REGION Network 15
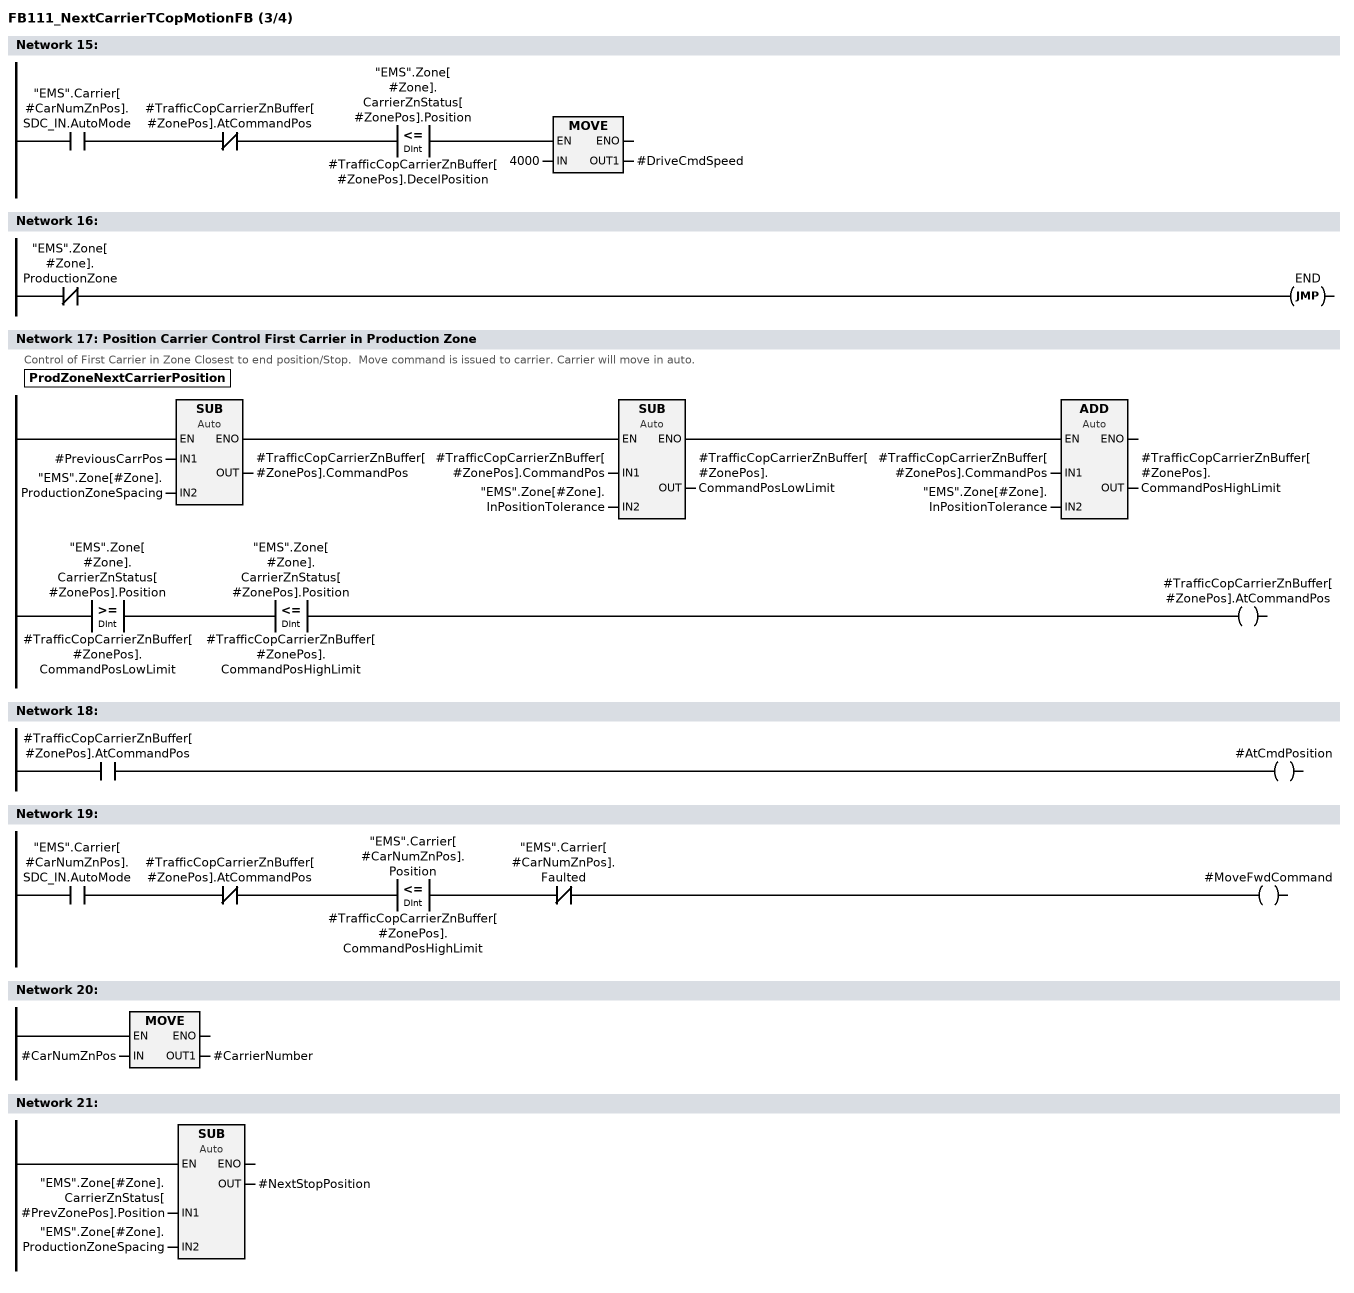
   RUNG wire#powerrail
      Contact( "EMS".Carrier[#CarNumZnPos].SDC_IN.AutoMode )
      I_Contact( #TrafficCopCarrierZnBuffer[#ZonePos].AtCommandPos )
      { S7_Templates := "SrcType := DInt" } LE_Contact(in1 := "EMS".Zone[#Zone].CarrierZnStatus[#ZonePos].Position, in2 := #TrafficCopCarrierZnBuffer[#ZonePos].DecelPosition)
      Move(in := 4000, out1 => #DriveCmdSpeed)
   END_RUNG
   // the same network as SCL:
   IF "EMS".Carrier[#CarNumZnPos].SDC_IN.AutoMode AND NOT #TrafficCopCarrierZnBuffer[#ZonePos].AtCommandPos AND ("EMS".Zone[#Zone].CarrierZnStatus[#ZonePos].Position <= #TrafficCopCarrierZnBuffer[#ZonePos].DecelPosition) THEN
       #DriveCmdSpeed := 4000;
   END_IF;
END_REGION

REGION Network 16
   RUNG wire#powerrail
      I_Contact( "EMS".Zone[#Zone].ProductionZone )
      JumpCoil( END )
   END_RUNG
   // the same network as SCL:
   IF NOT "EMS".Zone[#Zone].ProductionZone THEN GOTO END; END_IF;
END_REGION

REGION Network 17: Position Carrier Control First Carrier in Production Zone
   // Control of First Carrier in Zone Closest to end position/Stop.  Move command is issued to carrier. Carrier will move in auto.
   Label( ProdZoneNextCarrierPosition )
   RUNG wire#powerrail
      Sub(in1 := #PreviousCarrPos, in2 := "EMS".Zone[#Zone].ProductionZoneSpacing, out => #TrafficCopCarrierZnBuffer[#ZonePos].CommandPos)
      Sub(in1 := #TrafficCopCarrierZnBuffer[#ZonePos].CommandPos, in2 := "EMS".Zone[#Zone].InPositionTolerance, out => #TrafficCopCarrierZnBuffer[#ZonePos].CommandPosLowLimit)
      Add(in1 := #TrafficCopCarrierZnBuffer[#ZonePos].CommandPos, in2 := "EMS".Zone[#Zone].InPositionTolerance, out => #TrafficCopCarrierZnBuffer[#ZonePos].CommandPosHighLimit)
   END_RUNG
   RUNG wire#powerrail
      { S7_Templates := "SrcType := DInt" } GE_Contact(in1 := "EMS".Zone[#Zone].CarrierZnStatus[#ZonePos].Position, in2 := #TrafficCopCarrierZnBuffer[#ZonePos].CommandPosLowLimit)
      { S7_Templates := "SrcType := DInt" } LE_Contact(in1 := "EMS".Zone[#Zone].CarrierZnStatus[#ZonePos].Position, in2 := #TrafficCopCarrierZnBuffer[#ZonePos].CommandPosHighLimit)
      Coil( #TrafficCopCarrierZnBuffer[#ZonePos].AtCommandPos )
   END_RUNG
   // the same network as SCL:
   ProdZoneNextCarrierPosition:
   #TrafficCopCarrierZnBuffer[#ZonePos].CommandPos := #PreviousCarrPos - "EMS".Zone[#Zone].ProductionZoneSpacing;
   #TrafficCopCarrierZnBuffer[#ZonePos].CommandPosLowLimit := #TrafficCopCarrierZnBuffer[#ZonePos].CommandPos - "EMS".Zone[#Zone].InPositionTolerance;
   #TrafficCopCarrierZnBuffer[#ZonePos].CommandPosHighLimit := #TrafficCopCarrierZnBuffer[#ZonePos].CommandPos + "EMS".Zone[#Zone].InPositionTolerance;
   #TrafficCopCarrierZnBuffer[#ZonePos].AtCommandPos := ("EMS".Zone[#Zone].CarrierZnStatus[#ZonePos].Position >= #TrafficCopCarrierZnBuffer[#ZonePos].CommandPosLowLimit) AND ("EMS".Zone[#Zone].CarrierZnStatus[#ZonePos].Position <= #TrafficCopCarrierZnBuffer[#ZonePos].CommandPosHighLimit);
END_REGION

REGION Network 18
   RUNG wire#powerrail
      Contact( #TrafficCopCarrierZnBuffer[#ZonePos].AtCommandPos )
      Coil( #AtCmdPosition )
   END_RUNG
   // the same network as SCL:
   #AtCmdPosition := #TrafficCopCarrierZnBuffer[#ZonePos].AtCommandPos;
END_REGION

REGION Network 19
   RUNG wire#powerrail
      Contact( "EMS".Carrier[#CarNumZnPos].SDC_IN.AutoMode )
      I_Contact( #TrafficCopCarrierZnBuffer[#ZonePos].AtCommandPos )
      { S7_Templates := "SrcType := DInt" } LE_Contact(in1 := "EMS".Carrier[#CarNumZnPos].Position, in2 := #TrafficCopCarrierZnBuffer[#ZonePos].CommandPosHighLimit)
      I_Contact( "EMS".Carrier[#CarNumZnPos].Faulted )
      Coil( #MoveFwdCommand )
   END_RUNG
   // the same network as SCL:
   #MoveFwdCommand := "EMS".Carrier[#CarNumZnPos].SDC_IN.AutoMode AND NOT #TrafficCopCarrierZnBuffer[#ZonePos].AtCommandPos AND ("EMS".Carrier[#CarNumZnPos].Position <= #TrafficCopCarrierZnBuffer[#ZonePos].CommandPosHighLimit) AND NOT "EMS".Carrier[#CarNumZnPos].Faulted;
END_REGION

REGION Network 20
   RUNG wire#powerrail
      Move(in := #CarNumZnPos, out1 => #CarrierNumber)
   END_RUNG
   // the same network as SCL:
   #CarrierNumber := #CarNumZnPos;
END_REGION

REGION Network 21
   RUNG wire#powerrail
      Sub(in1 := "EMS".Zone[#Zone].CarrierZnStatus[#PrevZonePos].Position, in2 := "EMS".Zone[#Zone].ProductionZoneSpacing, out => #NextStopPosition)
   END_RUNG
   // the same network as SCL:
   #NextStopPosition := "EMS".Zone[#Zone].CarrierZnStatus[#PrevZonePos].Position - "EMS".Zone[#Zone].ProductionZoneSpacing;
END_REGION

REGION Network 22
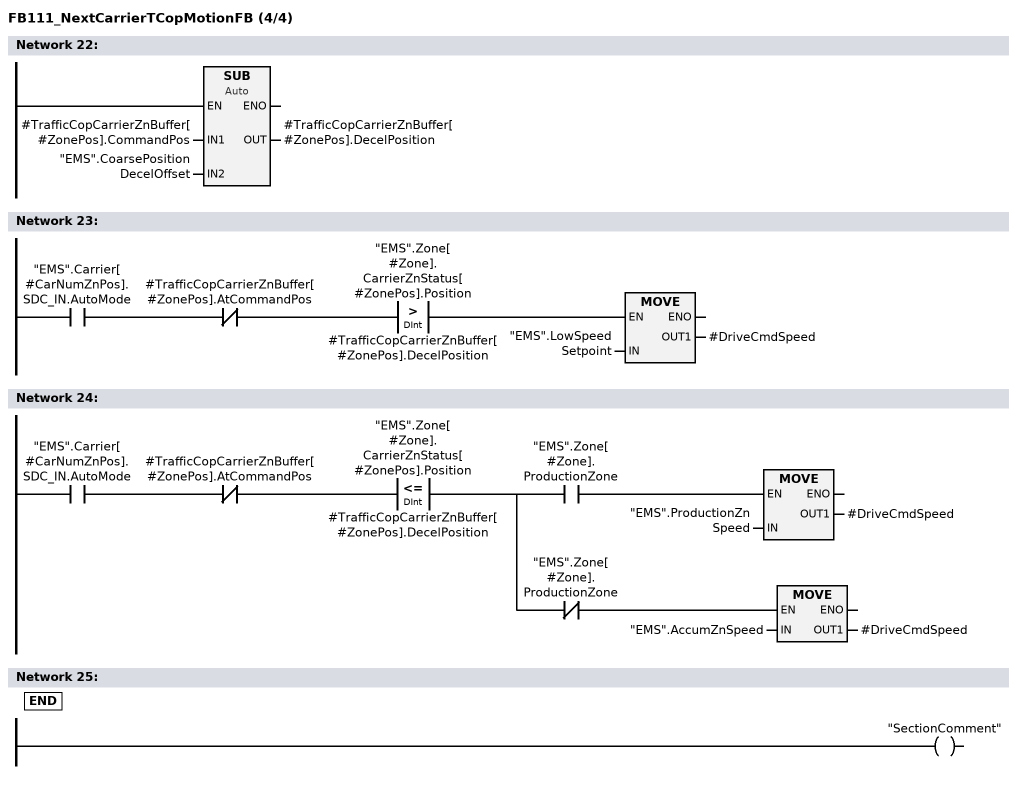
   RUNG wire#powerrail
      Sub(in1 := #TrafficCopCarrierZnBuffer[#ZonePos].CommandPos, in2 := "EMS".CoarsePositionDecelOffset, out => #TrafficCopCarrierZnBuffer[#ZonePos].DecelPosition)
   END_RUNG
   // the same network as SCL:
   #TrafficCopCarrierZnBuffer[#ZonePos].DecelPosition := #TrafficCopCarrierZnBuffer[#ZonePos].CommandPos - "EMS".CoarsePositionDecelOffset;
END_REGION

REGION Network 23
   RUNG wire#powerrail
      Contact( "EMS".Carrier[#CarNumZnPos].SDC_IN.AutoMode )
      I_Contact( #TrafficCopCarrierZnBuffer[#ZonePos].AtCommandPos )
      { S7_Templates := "SrcType := DInt" } GT_Contact(in1 := "EMS".Zone[#Zone].CarrierZnStatus[#ZonePos].Position, in2 := #TrafficCopCarrierZnBuffer[#ZonePos].DecelPosition)
      Move(in := "EMS".LowSpeedSetpoint, out1 => #DriveCmdSpeed)
   END_RUNG
   // the same network as SCL:
   IF "EMS".Carrier[#CarNumZnPos].SDC_IN.AutoMode AND NOT #TrafficCopCarrierZnBuffer[#ZonePos].AtCommandPos AND ("EMS".Zone[#Zone].CarrierZnStatus[#ZonePos].Position > #TrafficCopCarrierZnBuffer[#ZonePos].DecelPosition) THEN
       #DriveCmdSpeed := "EMS".LowSpeedSetpoint;
   END_IF;
END_REGION

REGION Network 24
   RUNG wire#powerrail
      Contact( "EMS".Carrier[#CarNumZnPos].SDC_IN.AutoMode )
      I_Contact( #TrafficCopCarrierZnBuffer[#ZonePos].AtCommandPos )
      { S7_Templates := "SrcType := DInt" } LE_Contact(in1 := "EMS".Zone[#Zone].CarrierZnStatus[#ZonePos].Position, in2 := #TrafficCopCarrierZnBuffer[#ZonePos].DecelPosition)
      wire#w1
      Contact( "EMS".Zone[#Zone].ProductionZone )
      Move(in := "EMS".ProductionZnSpeed, out1 => #DriveCmdSpeed)
   END_RUNG
   RUNG wire#w1
      I_Contact( "EMS".Zone[#Zone].ProductionZone )
      Move(in := "EMS".AccumZnSpeed, out1 => #DriveCmdSpeed)
   END_RUNG
   // the same network as SCL:
   #_w1 := "EMS".Carrier[#CarNumZnPos].SDC_IN.AutoMode AND NOT #TrafficCopCarrierZnBuffer[#ZonePos].AtCommandPos AND ("EMS".Zone[#Zone].CarrierZnStatus[#ZonePos].Position <= #TrafficCopCarrierZnBuffer[#ZonePos].DecelPosition);
   IF #_w1 AND "EMS".Zone[#Zone].ProductionZone THEN #DriveCmdSpeed := "EMS".ProductionZnSpeed; END_IF;
   IF #_w1 AND NOT "EMS".Zone[#Zone].ProductionZone THEN #DriveCmdSpeed := "EMS".AccumZnSpeed; END_IF;
END_REGION

REGION Network 25
   Label( END )
   RUNG wire#powerrail
      Coil( "SectionComment" )
   END_RUNG
   // the same network as SCL:
   END:
   "SectionComment" := TRUE;
END_REGION
END_FUNCTION_BLOCK

FUNCTION_BLOCK "FB112_Carrier"   // FB112, LAD
{ S7_Optimized_Access := 'TRUE' }
VERSION : 0.1
   VAR_INPUT
      Carrier : Int;
      EMS : "UDT_System";
      MoveFwd : Bool;
      SpeedSelect : Word;   // Speed Select 1=Slow 2=Normal
      CarrierFindArrayBufferiN : "UDT_Carrier";
      SDC_IN : "UDT_SDC_IN";
      DuplicateCarrierNumIn : Int;
      DuplicateCarrierFound : Bool;
      GapSpacingFault : Bool;
      FaultReset : Bool;
   END_VAR
   VAR_OUTPUT
      Zone : Int;
      ZonePos : Word;
      CarrierPositionEcho : DWord;
      CarrierNumberEcho : Word;
      DuplicateCarrierNumEcho : Word;
      CarrierNextStopPosEcho : Word;
      Faults : "UDT_SDCOutFaults";
      Faulted : Bool;
   END_VAR
   VAR
      CarrierMoveFwdSetup : Array[0..30] of Bool;
      MotionOffFaultTimer : IEC_TIMER;
      MotionOnFaultTimer : IEC_TIMER;
   END_VAR
BEGIN

REGION Network 1
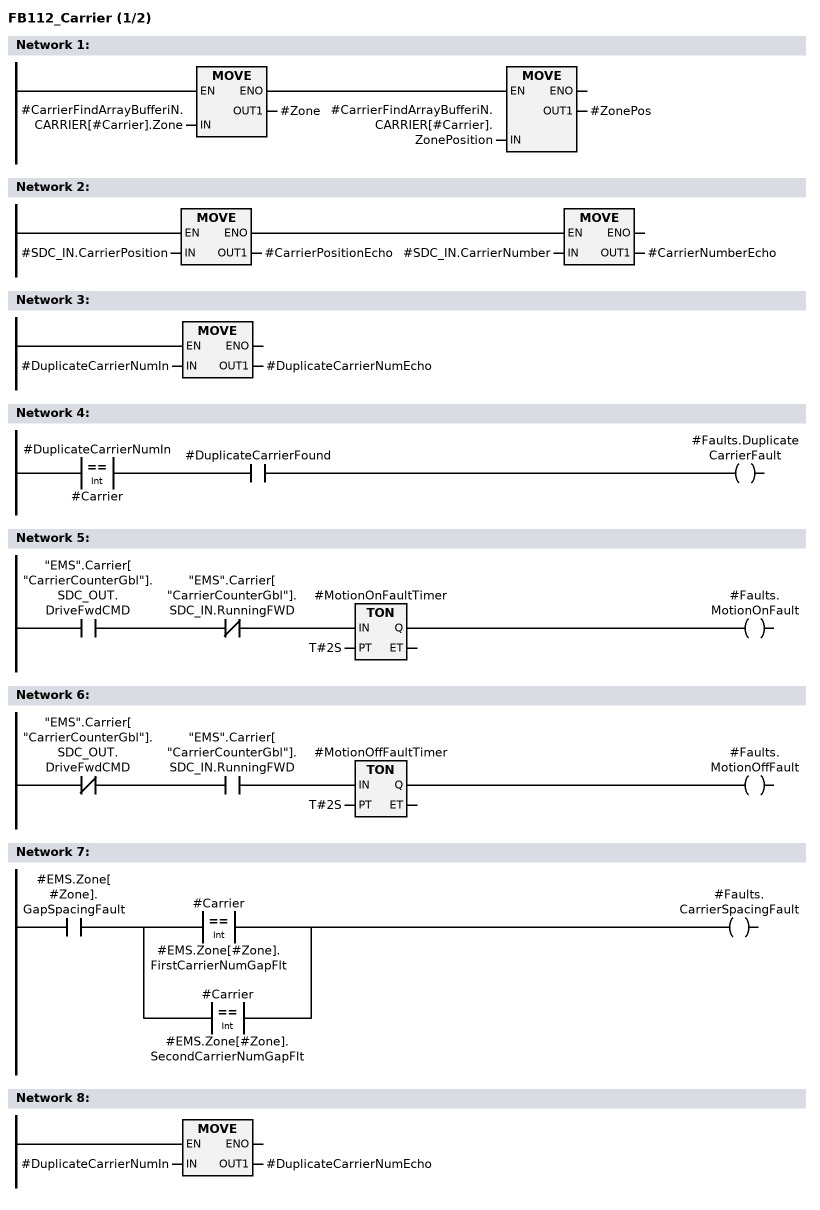
   RUNG wire#powerrail
      Move(in := #CarrierFindArrayBufferiN.CARRIER[#Carrier].Zone, out1 => #Zone)
      Move(in := #CarrierFindArrayBufferiN.CARRIER[#Carrier].ZonePosition, out1 => #ZonePos)
   END_RUNG
   // the same network as SCL:
   #Zone := #CarrierFindArrayBufferiN.CARRIER[#Carrier].Zone;
   #ZonePos := #CarrierFindArrayBufferiN.CARRIER[#Carrier].ZonePosition;
END_REGION

REGION Network 2
   RUNG wire#powerrail
      Move(in := #SDC_IN.CarrierPosition, out1 => #CarrierPositionEcho)
      Move(in := #SDC_IN.CarrierNumber, out1 => #CarrierNumberEcho)
   END_RUNG
   // the same network as SCL:
   #CarrierPositionEcho := #SDC_IN.CarrierPosition;
   #CarrierNumberEcho := #SDC_IN.CarrierNumber;
END_REGION

REGION Network 3
   RUNG wire#powerrail
      Move(in := #DuplicateCarrierNumIn, out1 => #DuplicateCarrierNumEcho)
   END_RUNG
   // the same network as SCL:
   #DuplicateCarrierNumEcho := #DuplicateCarrierNumIn;
END_REGION

REGION Network 4
   RUNG wire#powerrail
      { S7_Templates := "SrcType := Int" } EQ_Contact(in1 := #DuplicateCarrierNumIn, in2 := #Carrier)
      Contact( #DuplicateCarrierFound )
      Coil( #Faults.DuplicateCarrierFault )
   END_RUNG
   // the same network as SCL:
   #Faults.DuplicateCarrierFault := (#DuplicateCarrierNumIn = #Carrier) AND #DuplicateCarrierFound;
END_REGION

REGION Network 5
   #MotionOnFaultTimer.TON(IN := "EMS".Carrier["CarrierCounterGbl"].SDC_OUT.DriveFwdCMD AND NOT "EMS".Carrier["CarrierCounterGbl"].SDC_IN.RunningFWD,
                           PT := T#2S);
   #Faults.MotionOnFault := #MotionOnFaultTimer.Q;
END_REGION

REGION Network 6
   #MotionOffFaultTimer.TON(IN := NOT "EMS".Carrier["CarrierCounterGbl"].SDC_OUT.DriveFwdCMD AND "EMS".Carrier["CarrierCounterGbl"].SDC_IN.RunningFWD,
                           PT := T#2S);
   #Faults.MotionOffFault := #MotionOffFaultTimer.Q;
END_REGION

REGION Network 7
   RUNG wire#powerrail
      Contact( #EMS.Zone[#Zone].GapSpacingFault )
      wire#w1
      { S7_Templates := "SrcType := Int" } EQ_Contact(in1 := #Carrier, in2 := #EMS.Zone[#Zone].FirstCarrierNumGapFlt)
      wire#w2
      Coil( #Faults.CarrierSpacingFault )
   END_RUNG
   RUNG wire#w1
      { S7_Templates := "SrcType := Int" } EQ_Contact(in1 := #Carrier, in2 := #EMS.Zone[#Zone].SecondCarrierNumGapFlt)
   END_RUNG wire#w2
   // the same network as SCL:
   #Faults.CarrierSpacingFault := #EMS.Zone[#Zone].GapSpacingFault AND ((#Carrier = #EMS.Zone[#Zone].FirstCarrierNumGapFlt) OR (#Carrier = #EMS.Zone[#Zone].SecondCarrierNumGapFlt));
END_REGION

REGION Network 8
   RUNG wire#powerrail
      Move(in := #DuplicateCarrierNumIn, out1 => #DuplicateCarrierNumEcho)
   END_RUNG
   // the same network as SCL:
   #DuplicateCarrierNumEcho := #DuplicateCarrierNumIn;
END_REGION

REGION Network 9
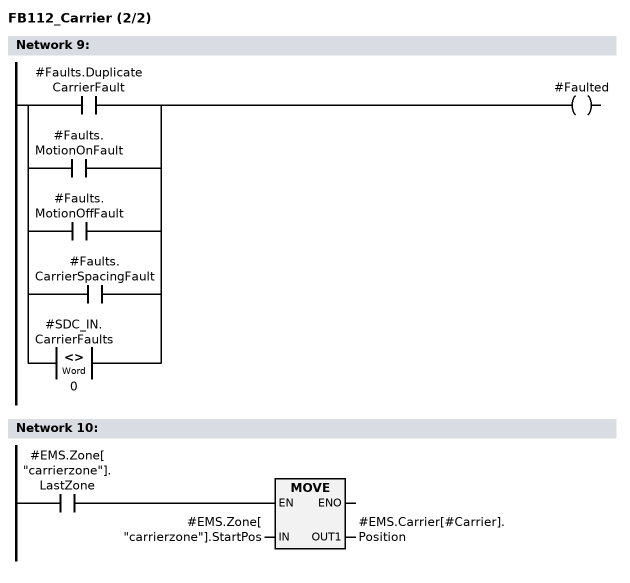
   RUNG wire#powerrail
      Contact( #Faults.DuplicateCarrierFault )
      wire#w1
      Coil( #Faulted )
   END_RUNG
   RUNG wire#powerrail
      Contact( #Faults.MotionOnFault )
   END_RUNG wire#w1
   RUNG wire#powerrail
      Contact( #Faults.MotionOffFault )
   END_RUNG wire#w1
   RUNG wire#powerrail
      Contact( #Faults.CarrierSpacingFault )
   END_RUNG wire#w1
   RUNG wire#powerrail
      { S7_Templates := "SrcType := Word" } NE_Contact(in1 := #SDC_IN.CarrierFaults, in2 := 0)
   END_RUNG wire#w1
   // the same network as SCL:
   #Faulted := #Faults.DuplicateCarrierFault OR #Faults.MotionOnFault OR #Faults.MotionOffFault OR #Faults.CarrierSpacingFault OR (#SDC_IN.CarrierFaults <> 0);
END_REGION

REGION Network 10
   RUNG wire#powerrail
      Contact( #EMS.Zone["carrierzone"].LastZone )
      Move(in := #EMS.Zone["carrierzone"].StartPos, out1 => #EMS.Carrier[#Carrier].Position)
   END_RUNG
   // the same network as SCL:
   IF #EMS.Zone["carrierzone"].LastZone THEN
       #EMS.Carrier[#Carrier].Position := #EMS.Zone["carrierzone"].StartPos;
   END_IF;
END_REGION
END_FUNCTION_BLOCK

FUNCTION_BLOCK "FB113_CarrierTrafficCop"   // FB113, LAD
{ S7_Optimized_Access := 'TRUE' }
VERSION : 0.1
   VAR_INPUT
      CarrierNumber : Word;
      ZonePos : Word;
   END_VAR
BEGIN
END_FUNCTION_BLOCK

FUNCTION_BLOCK "FB115_FB_Zone"   // FB115, LAD
{ S7_Optimized_Access := 'FALSE' }
VERSION : 0.1
   VAR_INPUT
      Zone : Int;
      Description : String[10];
      LastZone : Bool;
      MaxCarriers : Int;
      StartPos : DWord;
      EndPos : DWord;
      NextZone : Word;   // If Zone numbering is non sequential Next Zone Nu
      PreviousZone : Word;   // If Zone numbering is non sequential Previous Zone Nu
      SpeedZone : Bool;
      SpeedZoneStart : DWord;
      SpeedZoneEnd : DWord;
      AccumZone : Bool;
      AccumZnSpacing : Word;
      ProductionZone : Bool := false;
      ProductZoneSpacing : Word;
      FinePosStopZone : Bool;
      FineInPosTolerance : Word;
      FinePositionDecelOffset : Word;
      CoarseInPosTolerance : Word;
      CoarsePositionDecelOffset : Word;
      NextCarrierClrHighSpeed : Word;
      StopControlFromEMS01 : "UDT_StopControlFromEMS01";
   END_VAR
   VAR_OUTPUT
      ZoneEcho : Word;
      LastZoneEcho : Bool;
      ZoneFull : Bool;
      ZoneLengthEcho : Word;
      DescriptionEcho : String[10];
      StartPosEcho : DWord;
      EndPosEcho : DWord;
      SpeedZoneEcho : Bool;
      SpeedZoneStartEcho : DWord;
      SpeedZoneEndEcho : DWord;
      AccumZoneEcho : Bool;
      AccumSpacingEcho : Word;
      ProductionZoneEcho : Bool;
      ProdZoneSpacingEcho : Word;
      CarrierInPosToleranceEcho : Word;
      NextCarrierClrHighSpeedEcho : Word;
      MaxCarriersEcho : Word;
      ClearToEnterEcho : Bool;
      ClearZoneStartEcho : Bool;
      ClearZoneEcho : Bool;
      ZoneCarrierStatsArray : Array[0..60] of "UDT_ZoneCarrierStatus";
      FinePosStopZoneEcho : Bool;
      FineInPosToleranceEcho : Word;
      FinePositionDecelEcho : Word;
      CoarsePositionDecelEcho : Word;
      CoarseInPosToleranceEcho : Word;
      PreviosZoneEcho : Word;
      NextZoneEcho : Word;
      CarrierAtStop : Bool;
      CarrierNumAtStop : Word;
      HMIZonePositionsEcho : Array[1..20] of "UDT_HMIZonePositions";
      ClearOfStopPos : DWord;
      StopStatusToEMS01 : "UDT_StopStatusToEMS01";
   END_VAR
   VAR_TEMP
      HMIZonePositions : Array[1..20] of "UDT_HMIZonePositions";
      carrierstatusdn : Bool;
      resettemp : Bool;
      resettemp2 : Bool;
      sortdonetemp : Bool;
      ZonePosSpacing : Word;
      ZoneLengthTemp : UDInt;
   END_VAR
BEGIN

REGION Network 1
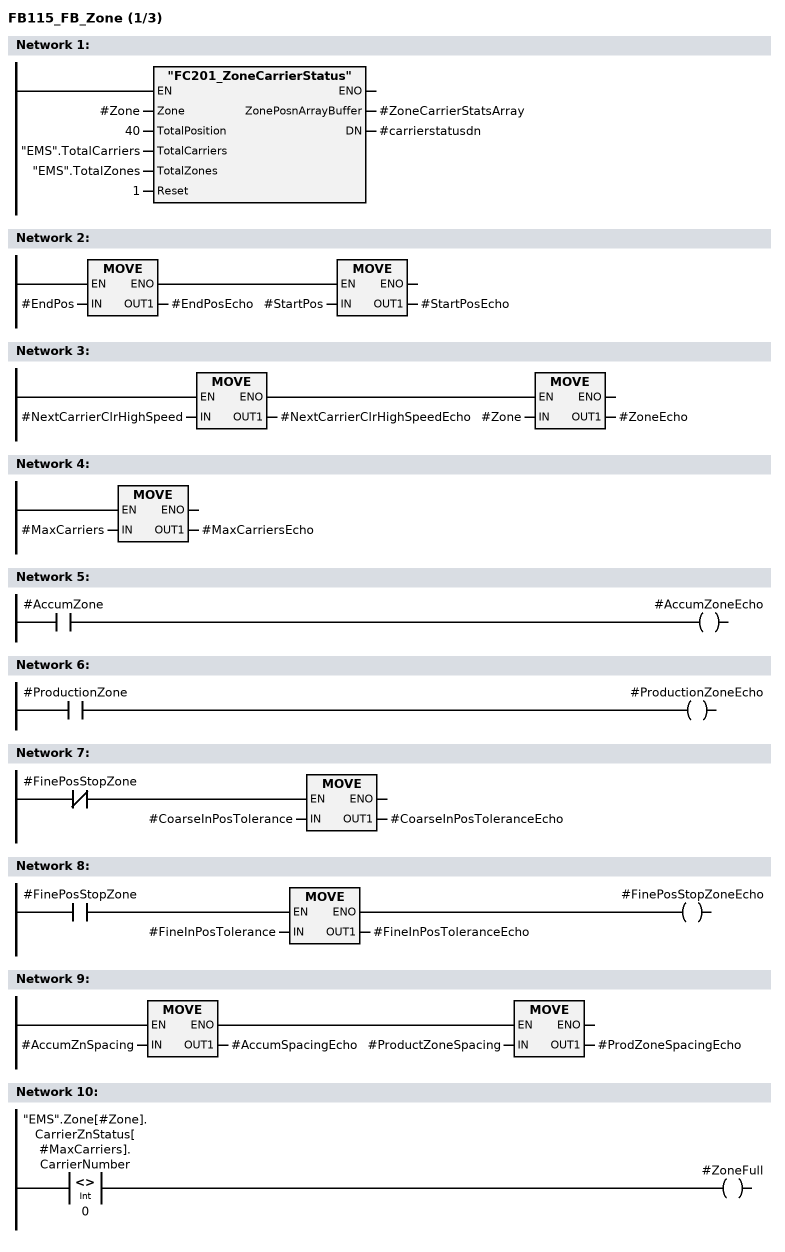
   RUNG wire#powerrail
      "FC201_ZoneCarrierStatus"(Zone := #Zone, TotalPosition := 40, TotalCarriers := "EMS".TotalCarriers, TotalZones := "EMS".TotalZones, Reset := 1, ZonePosnArrayBuffer => #ZoneCarrierStatsArray, DN => #carrierstatusdn)
   END_RUNG
   // the same network as SCL:
   "FC201_ZoneCarrierStatus"(Zone := #Zone,
                           TotalPosition := 40,
                           TotalCarriers := "EMS".TotalCarriers,
                           TotalZones := "EMS".TotalZones,
                           Reset := 1,
                           ZonePosnArrayBuffer => #ZoneCarrierStatsArray,
                           DN => #carrierstatusdn);
END_REGION

REGION Network 2
   RUNG wire#powerrail
      Move(in := #EndPos, out1 => #EndPosEcho)
      Move(in := #StartPos, out1 => #StartPosEcho)
   END_RUNG
   // the same network as SCL:
   #EndPosEcho := #EndPos;
   #StartPosEcho := #StartPos;
END_REGION

REGION Network 3
   RUNG wire#powerrail
      Move(in := #NextCarrierClrHighSpeed, out1 => #NextCarrierClrHighSpeedEcho)
      Move(in := #Zone, out1 => #ZoneEcho)
   END_RUNG
   // the same network as SCL:
   #NextCarrierClrHighSpeedEcho := #NextCarrierClrHighSpeed;
   #ZoneEcho := #Zone;
END_REGION

REGION Network 4
   RUNG wire#powerrail
      Move(in := #MaxCarriers, out1 => #MaxCarriersEcho)
   END_RUNG
   // the same network as SCL:
   #MaxCarriersEcho := #MaxCarriers;
END_REGION

REGION Network 5
   RUNG wire#powerrail
      Contact( #AccumZone )
      Coil( #AccumZoneEcho )
   END_RUNG
   // the same network as SCL:
   #AccumZoneEcho := #AccumZone;
END_REGION

REGION Network 6
   RUNG wire#powerrail
      Contact( #ProductionZone )
      Coil( #ProductionZoneEcho )
   END_RUNG
   // the same network as SCL:
   #ProductionZoneEcho := #ProductionZone;
END_REGION

REGION Network 7
   RUNG wire#powerrail
      I_Contact( #FinePosStopZone )
      Move(in := #CoarseInPosTolerance, out1 => #CoarseInPosToleranceEcho)
   END_RUNG
   // the same network as SCL:
   IF NOT #FinePosStopZone THEN #CoarseInPosToleranceEcho := #CoarseInPosTolerance; END_IF;
END_REGION

REGION Network 8
   RUNG wire#powerrail
      Contact( #FinePosStopZone )
      Move(in := #FineInPosTolerance, out1 => #FineInPosToleranceEcho)
      Coil( #FinePosStopZoneEcho )
   END_RUNG
   // the same network as SCL:
   IF #FinePosStopZone THEN #FineInPosToleranceEcho := #FineInPosTolerance; END_IF;
   #FinePosStopZoneEcho := #FinePosStopZone;
END_REGION

REGION Network 9
   RUNG wire#powerrail
      Move(in := #AccumZnSpacing, out1 => #AccumSpacingEcho)
      Move(in := #ProductZoneSpacing, out1 => #ProdZoneSpacingEcho)
   END_RUNG
   // the same network as SCL:
   #AccumSpacingEcho := #AccumZnSpacing;
   #ProdZoneSpacingEcho := #ProductZoneSpacing;
END_REGION

REGION Network 10
   RUNG wire#powerrail
      { S7_Templates := "SrcType := Int" } NE_Contact(in1 := "EMS".Zone[#Zone].CarrierZnStatus[#MaxCarriers].CarrierNumber, in2 := 0)
      Coil( #ZoneFull )
   END_RUNG
   // the same network as SCL:
   #ZoneFull := "EMS".Zone[#Zone].CarrierZnStatus[#MaxCarriers].CarrierNumber <> 0;
END_REGION

REGION Network 11
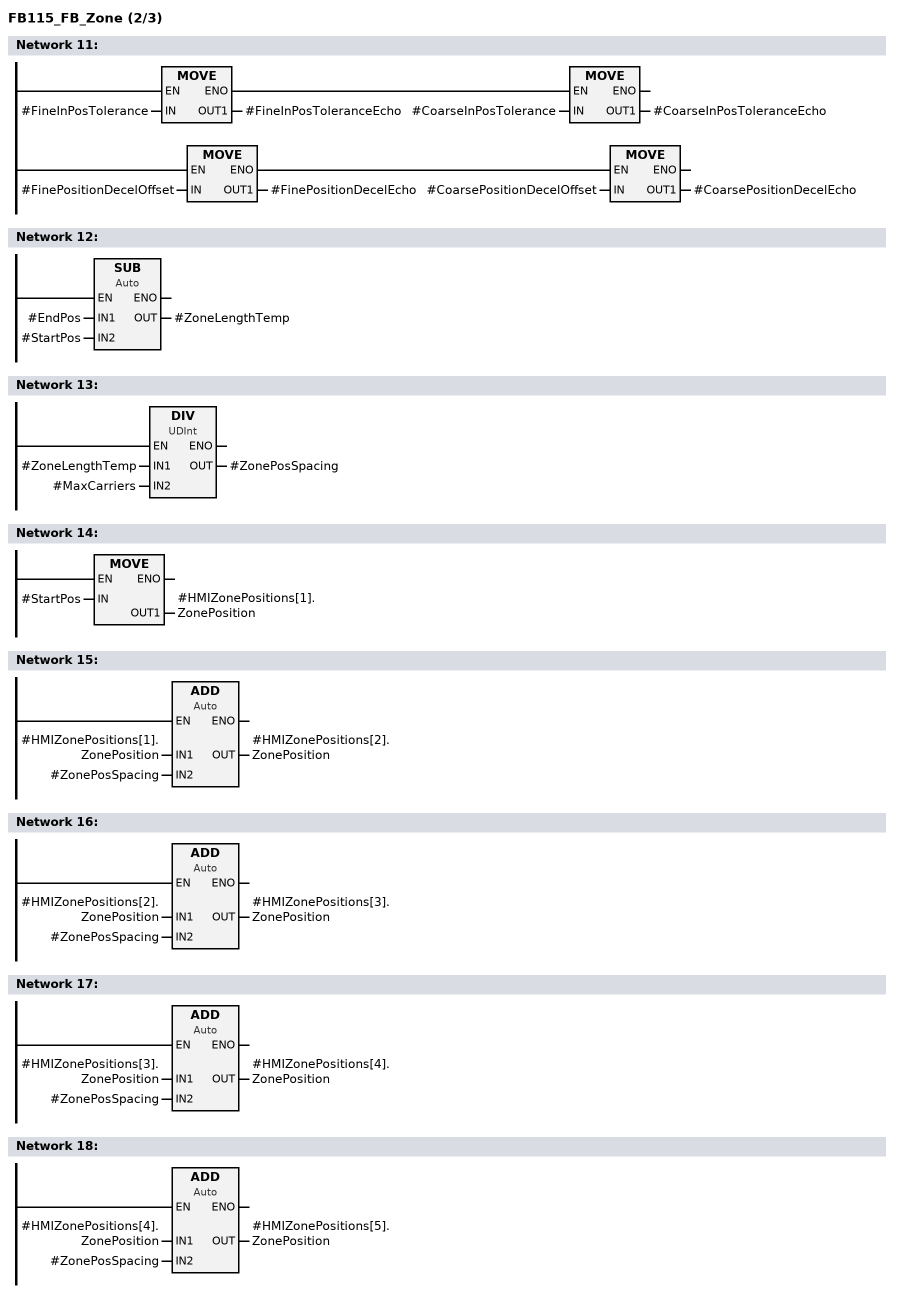
   RUNG wire#powerrail
      Move(in := #FineInPosTolerance, out1 => #FineInPosToleranceEcho)
      Move(in := #CoarseInPosTolerance, out1 => #CoarseInPosToleranceEcho)
   END_RUNG
   RUNG wire#powerrail
      Move(in := #FinePositionDecelOffset, out1 => #FinePositionDecelEcho)
      Move(in := #CoarsePositionDecelOffset, out1 => #CoarsePositionDecelEcho)
   END_RUNG
   // the same network as SCL:
   #FineInPosToleranceEcho := #FineInPosTolerance;
   #CoarseInPosToleranceEcho := #CoarseInPosTolerance;
   #FinePositionDecelEcho := #FinePositionDecelOffset;
   #CoarsePositionDecelEcho := #CoarsePositionDecelOffset;
END_REGION

REGION Network 12
   RUNG wire#powerrail
      Sub(in1 := #EndPos, in2 := #StartPos, out => #ZoneLengthTemp)
   END_RUNG
   // the same network as SCL:
   #ZoneLengthTemp := #EndPos - #StartPos;
END_REGION

REGION Network 13
   RUNG wire#powerrail
      { S7_Templates := "SrcType := UDInt" } Div(in1 := #ZoneLengthTemp, in2 := #MaxCarriers, out => #ZonePosSpacing)
   END_RUNG
   // the same network as SCL:
   #ZonePosSpacing := #ZoneLengthTemp / #MaxCarriers;
END_REGION

REGION Network 14
   RUNG wire#powerrail
      Move(in := #StartPos, out1 => #HMIZonePositions[1].ZonePosition)
   END_RUNG
   // the same network as SCL:
   #HMIZonePositions[1].ZonePosition := #StartPos;
END_REGION

REGION Network 15
   RUNG wire#powerrail
      Add(in1 := #HMIZonePositions[1].ZonePosition, in2 := #ZonePosSpacing, out => #HMIZonePositions[2].ZonePosition)
   END_RUNG
   // the same network as SCL:
   #HMIZonePositions[2].ZonePosition := #HMIZonePositions[1].ZonePosition + #ZonePosSpacing;
END_REGION

REGION Network 16
   RUNG wire#powerrail
      Add(in1 := #HMIZonePositions[2].ZonePosition, in2 := #ZonePosSpacing, out => #HMIZonePositions[3].ZonePosition)
   END_RUNG
   // the same network as SCL:
   #HMIZonePositions[3].ZonePosition := #HMIZonePositions[2].ZonePosition + #ZonePosSpacing;
END_REGION

REGION Network 17
   RUNG wire#powerrail
      Add(in1 := #HMIZonePositions[3].ZonePosition, in2 := #ZonePosSpacing, out => #HMIZonePositions[4].ZonePosition)
   END_RUNG
   // the same network as SCL:
   #HMIZonePositions[4].ZonePosition := #HMIZonePositions[3].ZonePosition + #ZonePosSpacing;
END_REGION

REGION Network 18
   RUNG wire#powerrail
      Add(in1 := #HMIZonePositions[4].ZonePosition, in2 := #ZonePosSpacing, out => #HMIZonePositions[5].ZonePosition)
   END_RUNG
   // the same network as SCL:
   #HMIZonePositions[5].ZonePosition := #HMIZonePositions[4].ZonePosition + #ZonePosSpacing;
END_REGION

REGION Network 19
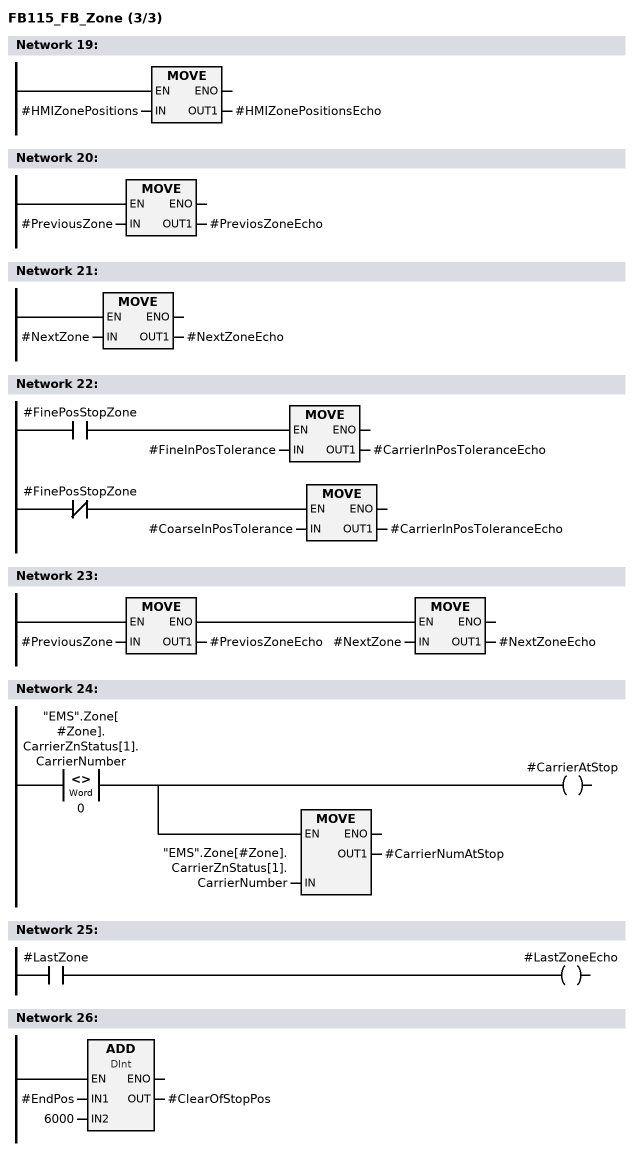
   RUNG wire#powerrail
      Move(in := #HMIZonePositions, out1 => #HMIZonePositionsEcho)
   END_RUNG
   // the same network as SCL:
   #HMIZonePositionsEcho := #HMIZonePositions;
END_REGION

REGION Network 20
   RUNG wire#powerrail
      Move(in := #PreviousZone, out1 => #PreviosZoneEcho)
   END_RUNG
   // the same network as SCL:
   #PreviosZoneEcho := #PreviousZone;
END_REGION

REGION Network 21
   RUNG wire#powerrail
      Move(in := #NextZone, out1 => #NextZoneEcho)
   END_RUNG
   // the same network as SCL:
   #NextZoneEcho := #NextZone;
END_REGION

REGION Network 22
   RUNG wire#powerrail
      Contact( #FinePosStopZone )
      Move(in := #FineInPosTolerance, out1 => #CarrierInPosToleranceEcho)
   END_RUNG
   RUNG wire#powerrail
      I_Contact( #FinePosStopZone )
      Move(in := #CoarseInPosTolerance, out1 => #CarrierInPosToleranceEcho)
   END_RUNG
   // the same network as SCL:
   IF #FinePosStopZone THEN #CarrierInPosToleranceEcho := #FineInPosTolerance; END_IF;
   IF NOT #FinePosStopZone THEN #CarrierInPosToleranceEcho := #CoarseInPosTolerance; END_IF;
END_REGION

REGION Network 23
   RUNG wire#powerrail
      Move(in := #PreviousZone, out1 => #PreviosZoneEcho)
      Move(in := #NextZone, out1 => #NextZoneEcho)
   END_RUNG
   // the same network as SCL:
   #PreviosZoneEcho := #PreviousZone;
   #NextZoneEcho := #NextZone;
END_REGION

REGION Network 24
   RUNG wire#powerrail
      { S7_Templates := "SrcType := Word" } NE_Contact(in1 := "EMS".Zone[#Zone].CarrierZnStatus[1].CarrierNumber, in2 := 0)
      wire#w1
      Coil( #CarrierAtStop )
   END_RUNG
   RUNG wire#w1
      Move(in := "EMS".Zone[#Zone].CarrierZnStatus[1].CarrierNumber, out1 => #CarrierNumAtStop)
   END_RUNG
   // the same network as SCL:
   #CarrierAtStop := "EMS".Zone[#Zone].CarrierZnStatus[1].CarrierNumber <> 0;
   IF #CarrierAtStop THEN #CarrierNumAtStop := "EMS".Zone[#Zone].CarrierZnStatus[1].CarrierNumber; END_IF;
END_REGION

REGION Network 25
   RUNG wire#powerrail
      Contact( #LastZone )
      Coil( #LastZoneEcho )
   END_RUNG
   // the same network as SCL:
   #LastZoneEcho := #LastZone;
END_REGION

REGION Network 26
   RUNG wire#powerrail
      { S7_Templates := "SrcType := DInt" } Add(in1 := #EndPos, in2 := 6000, out => #ClearOfStopPos)
   END_RUNG
   // the same network as SCL:
   #ClearOfStopPos := #EndPos + 6000;
END_REGION
END_FUNCTION_BLOCK

FUNCTION_BLOCK "FB116_FB_ZonePositionArrayTrafficCop"   // FB116, LAD
{ S7_Optimized_Access := 'FALSE' }
VERSION : 0.1
   VAR_INPUT
      Zone : Int := 1;
      CarrierZnArrayPos : Int;
   END_VAR
   VAR_OUTPUT
      MoveFwd : Bool;
      Speed : Word;
      TCZnPosnArray : "UDT_TrafficCopZoneStructure";
   END_VAR
   VAR
      CarNumZnPos : Array[0..99] of Int;
      TrafficCopCarrierZnBufferOut : Array[0..30] of "UDT_TrafficCop";
      "Zn-Pos2CarrierNumTemp" : Int;
      Zone1TrafficCopStructure : Struct
         CommandPosition : Word;
         InPositionTolerance : Word;
         CommandPositionUpperLimit : Word;
         CommandPositionLowerLimit : Word;
         AtCommandPos : Bool;
      END_STRUCT;
      SectionComment : Bool;
      NextCarrierZnArrayPos : Int;
   END_VAR
BEGIN

REGION Network 1: Section Comment-Section Logic for Current Carrier number in Position 1 thru Max Carrier in Zone Position Array
   // Section Logic for Current Carrier number in Position 1 - Max Carrier in Zone Position Array
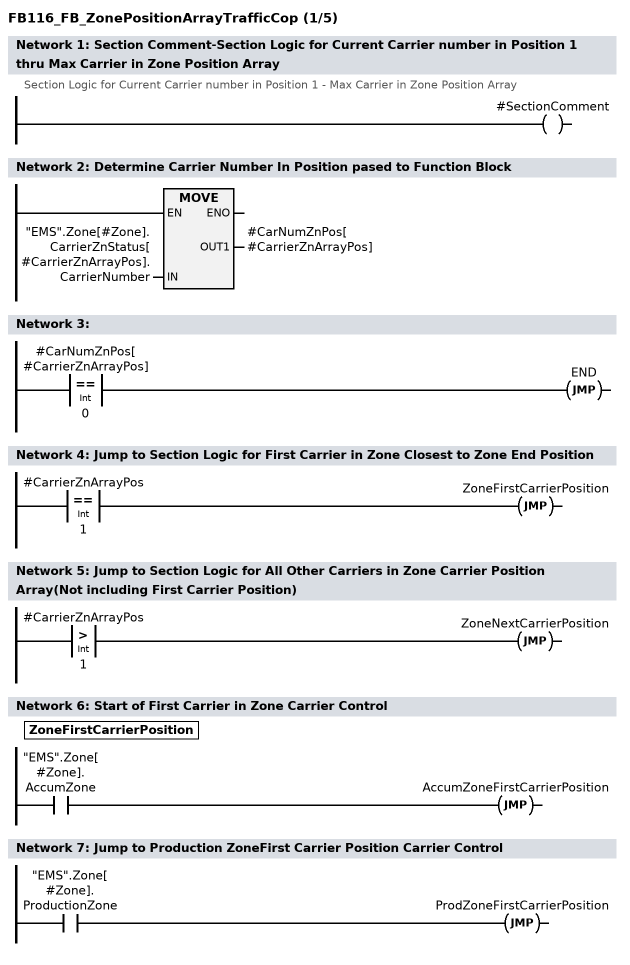
   RUNG wire#powerrail
      Coil( #SectionComment )
   END_RUNG
   // the same network as SCL:
   #SectionComment := TRUE;
END_REGION

REGION Network 2: Determine Carrier Number In Position pased to Function Block
   RUNG wire#powerrail
      Move(in := "EMS".Zone[#Zone].CarrierZnStatus[#CarrierZnArrayPos].CarrierNumber, out1 => #CarNumZnPos[#CarrierZnArrayPos])
   END_RUNG
   // the same network as SCL:
   #CarNumZnPos[#CarrierZnArrayPos] := "EMS".Zone[#Zone].CarrierZnStatus[#CarrierZnArrayPos].CarrierNumber;
END_REGION

REGION Network 3
   RUNG wire#powerrail
      { S7_Templates := "SrcType := Int" } EQ_Contact(in1 := #CarNumZnPos[#CarrierZnArrayPos], in2 := 0)
      JumpCoil( END )
   END_RUNG
   // the same network as SCL:
   IF #CarNumZnPos[#CarrierZnArrayPos] = 0 THEN GOTO END; END_IF;
END_REGION

REGION Network 4: Jump to Section Logic for First Carrier in Zone Closest to Zone End Position
   RUNG wire#powerrail
      { S7_Templates := "SrcType := Int" } EQ_Contact(in1 := #CarrierZnArrayPos, in2 := 1)
      JumpCoil( ZoneFirstCarrierPosition )
   END_RUNG
   // the same network as SCL:
   IF #CarrierZnArrayPos = 1 THEN GOTO ZoneFirstCarrierPosition; END_IF;
END_REGION

REGION Network 5: Jump to Section Logic for All Other Carriers in Zone Carrier Position Array(Not including First Carrier Position)
   RUNG wire#powerrail
      { S7_Templates := "SrcType := Int" } GT_Contact(in1 := #CarrierZnArrayPos, in2 := 1)
      JumpCoil( ZoneNextCarrierPosition )
   END_RUNG
   // the same network as SCL:
   IF #CarrierZnArrayPos > 1 THEN GOTO ZoneNextCarrierPosition; END_IF;
END_REGION

REGION Network 6: Start of First Carrier in Zone Carrier Control
   Label( ZoneFirstCarrierPosition )
   RUNG wire#powerrail
      Contact( "EMS".Zone[#Zone].AccumZone )
      JumpCoil( AccumZoneFirstCarrierPosition )
   END_RUNG
   // the same network as SCL:
   ZoneFirstCarrierPosition:
   IF "EMS".Zone[#Zone].AccumZone THEN GOTO AccumZoneFirstCarrierPosition; END_IF;
END_REGION

REGION Network 7: Jump to Production ZoneFirst Carrier Position Carrier Control
   RUNG wire#powerrail
      Contact( "EMS".Zone[#Zone].ProductionZone )
      JumpCoil( ProdZoneFirstCarrierPosition )
   END_RUNG
   // the same network as SCL:
   IF "EMS".Zone[#Zone].ProductionZone THEN GOTO ProdZoneFirstCarrierPosition; END_IF;
END_REGION

REGION Network 8: Position Carrier Control First Carrier in Accumulation Zone
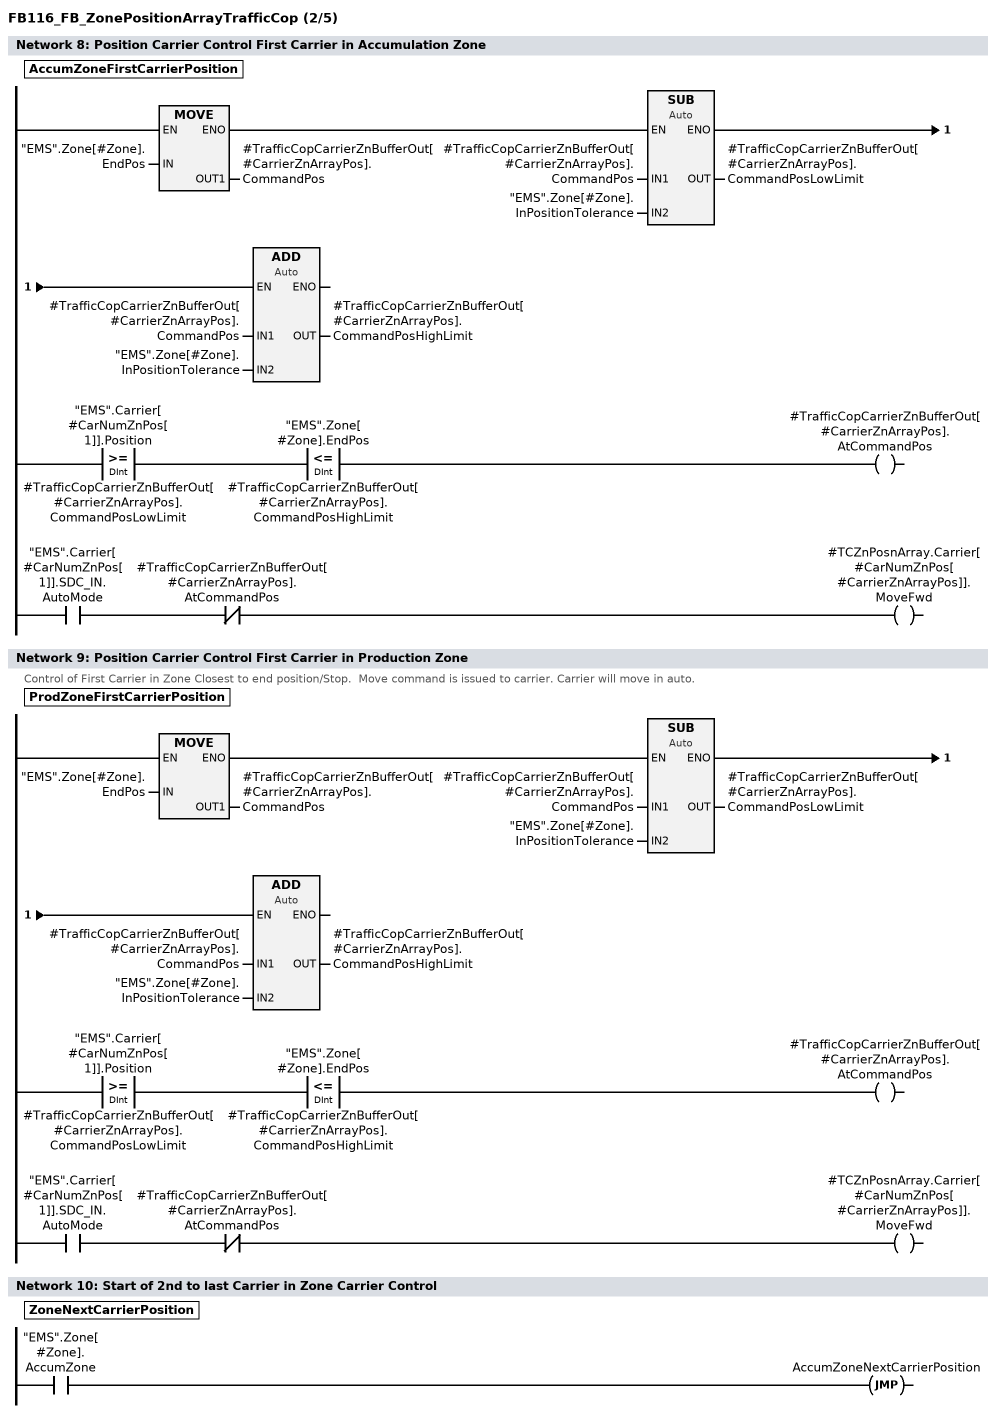
   Label( AccumZoneFirstCarrierPosition )
   RUNG wire#powerrail
      Move(in := "EMS".Zone[#Zone].EndPos, out1 => #TrafficCopCarrierZnBufferOut[#CarrierZnArrayPos].CommandPos)
      Sub(in1 := #TrafficCopCarrierZnBufferOut[#CarrierZnArrayPos].CommandPos, in2 := "EMS".Zone[#Zone].InPositionTolerance, out => #TrafficCopCarrierZnBufferOut[#CarrierZnArrayPos].CommandPosLowLimit)
      Add(in1 := #TrafficCopCarrierZnBufferOut[#CarrierZnArrayPos].CommandPos, in2 := "EMS".Zone[#Zone].InPositionTolerance, out => #TrafficCopCarrierZnBufferOut[#CarrierZnArrayPos].CommandPosHighLimit)
   END_RUNG
   RUNG wire#powerrail
      { S7_Templates := "SrcType := DInt" } GE_Contact(in1 := "EMS".Carrier[#CarNumZnPos[1]].Position, in2 := #TrafficCopCarrierZnBufferOut[#CarrierZnArrayPos].CommandPosLowLimit)
      { S7_Templates := "SrcType := DInt" } LE_Contact(in1 := "EMS".Zone[#Zone].EndPos, in2 := #TrafficCopCarrierZnBufferOut[#CarrierZnArrayPos].CommandPosHighLimit)
      Coil( #TrafficCopCarrierZnBufferOut[#CarrierZnArrayPos].AtCommandPos )
   END_RUNG
   RUNG wire#powerrail
      Contact( "EMS".Carrier[#CarNumZnPos[1]].SDC_IN.AutoMode )
      I_Contact( #TrafficCopCarrierZnBufferOut[#CarrierZnArrayPos].AtCommandPos )
      Coil( #TCZnPosnArray.Carrier[#CarNumZnPos[#CarrierZnArrayPos]].MoveFwd )
   END_RUNG
   // the same network as SCL:
   AccumZoneFirstCarrierPosition:
   #TrafficCopCarrierZnBufferOut[#CarrierZnArrayPos].CommandPos := "EMS".Zone[#Zone].EndPos;
   #TrafficCopCarrierZnBufferOut[#CarrierZnArrayPos].CommandPosLowLimit := #TrafficCopCarrierZnBufferOut[#CarrierZnArrayPos].CommandPos - "EMS".Zone[#Zone].InPositionTolerance;
   #TrafficCopCarrierZnBufferOut[#CarrierZnArrayPos].CommandPosHighLimit := #TrafficCopCarrierZnBufferOut[#CarrierZnArrayPos].CommandPos + "EMS".Zone[#Zone].InPositionTolerance;
   #TrafficCopCarrierZnBufferOut[#CarrierZnArrayPos].AtCommandPos := ("EMS".Carrier[#CarNumZnPos[1]].Position >= #TrafficCopCarrierZnBufferOut[#CarrierZnArrayPos].CommandPosLowLimit) AND ("EMS".Zone[#Zone].EndPos <= #TrafficCopCarrierZnBufferOut[#CarrierZnArrayPos].CommandPosHighLimit);
   #TCZnPosnArray.Carrier[#CarNumZnPos[#CarrierZnArrayPos]].MoveFwd := "EMS".Carrier[#CarNumZnPos[1]].SDC_IN.AutoMode AND NOT #TrafficCopCarrierZnBufferOut[#CarrierZnArrayPos].AtCommandPos;
END_REGION
